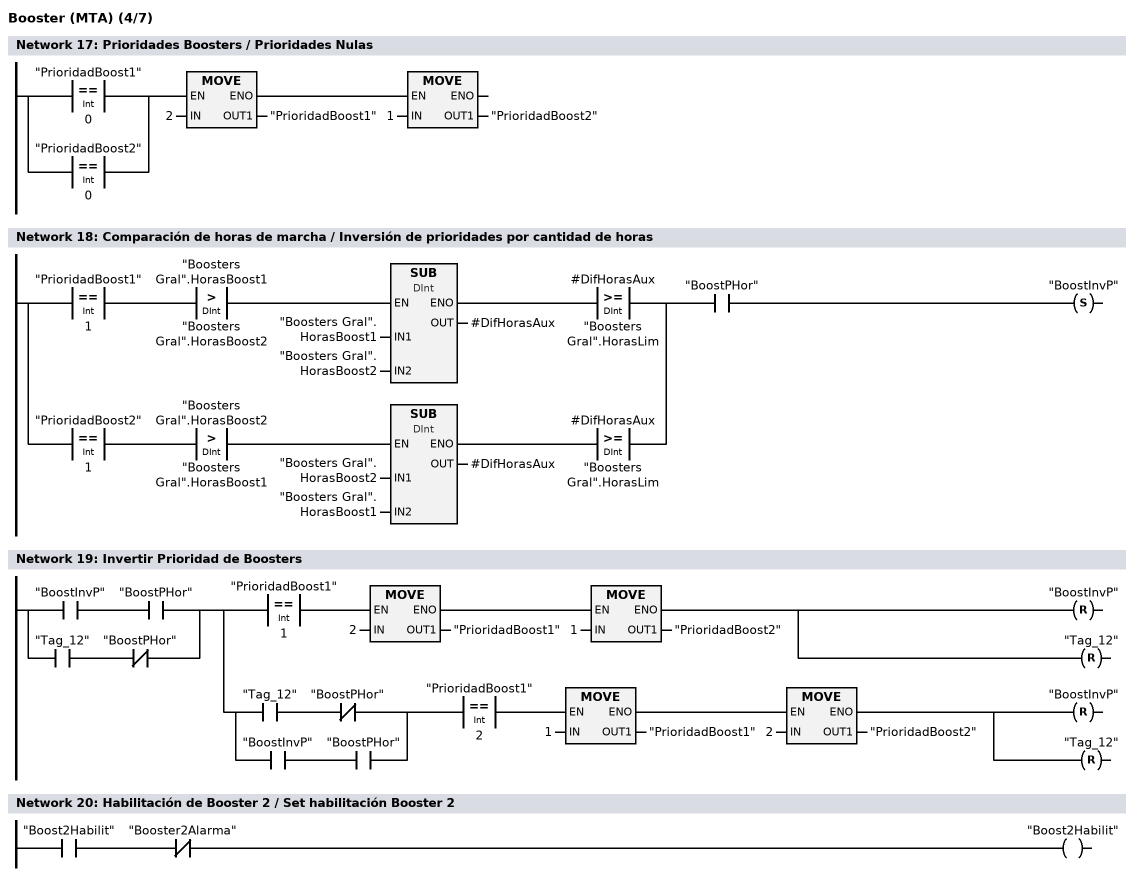
   RUNG wire#powerrail
      { S7_Templates := "SrcType := Int" } EQ_Contact(in1 := "PrioridadBoost1", in2 := 0)
      wire#w1
      { S7_GenerateENO := "TRUE" } Move(in := 2, out1 => "PrioridadBoost1")
      { S7_GenerateENO := "TRUE" } Move(in := 1, out1 => "PrioridadBoost2")
   END_RUNG
   RUNG wire#powerrail
      { S7_Templates := "SrcType := Int" } EQ_Contact(in1 := "PrioridadBoost2", in2 := 0)
   END_RUNG wire#w1
   // the same network as SCL:
   // ENO of a box is taken as its EN; it also drops when the box reports an error
   #_w1 := ("PrioridadBoost1" = 0) OR ("PrioridadBoost2" = 0);
   IF #_w1 THEN
       "PrioridadBoost1" := 2;
       "PrioridadBoost2" := 1;
   END_IF;
END_REGION

REGION Network 18: Comparación de horas de marcha / Inversión de prioridades por cantidad de horas
   RUNG wire#powerrail
      { S7_Templates := "SrcType := Int" } EQ_Contact(in1 := "PrioridadBoost1", in2 := 1)
      { S7_Templates := "SrcType := DInt" } GT_Contact(in1 := "Boosters Gral".HorasBoost1, in2 := "Boosters Gral".HorasBoost2)
      { S7_Templates := "SrcType := DInt"; S7_GenerateENO := "TRUE" } Sub(in1 := "Boosters Gral".HorasBoost1, in2 := "Boosters Gral".HorasBoost2, out => #DifHorasAux)
      { S7_Templates := "SrcType := DInt" } GE_Contact(in1 := #DifHorasAux, in2 := "Boosters Gral".HorasLim)
      wire#w1
      Contact( "BoostPHor" )
      S_Coil( "BoostInvP" )
   END_RUNG
   RUNG wire#powerrail
      { S7_Templates := "SrcType := Int" } EQ_Contact(in1 := "PrioridadBoost2", in2 := 1)
      { S7_Templates := "SrcType := DInt" } GT_Contact(in1 := "Boosters Gral".HorasBoost2, in2 := "Boosters Gral".HorasBoost1)
      { S7_Templates := "SrcType := DInt"; S7_GenerateENO := "TRUE" } Sub(in1 := "Boosters Gral".HorasBoost2, in2 := "Boosters Gral".HorasBoost1, out => #DifHorasAux)
      { S7_Templates := "SrcType := DInt" } GE_Contact(in1 := #DifHorasAux, in2 := "Boosters Gral".HorasLim)
   END_RUNG wire#w1
   // the same network as SCL:
   // ENO of a box is taken as its EN; it also drops when the box reports an error
   #_w1 := ("PrioridadBoost1" = 1) AND ("Boosters Gral".HorasBoost1 > "Boosters Gral".HorasBoost2);
   IF #_w1 THEN #DifHorasAux := "Boosters Gral".HorasBoost1 - "Boosters Gral".HorasBoost2; END_IF;
   #_w2 := ("PrioridadBoost2" = 1) AND ("Boosters Gral".HorasBoost2 > "Boosters Gral".HorasBoost1);
   #_w3 := #_w1 AND (#DifHorasAux >= "Boosters Gral".HorasLim);
   IF #_w2 THEN #DifHorasAux := "Boosters Gral".HorasBoost2 - "Boosters Gral".HorasBoost1; END_IF;
   IF (#_w3 OR (#_w2 AND (#DifHorasAux >= "Boosters Gral".HorasLim))) AND "BoostPHor" THEN
       "BoostInvP" := TRUE;
   END_IF;
END_REGION

REGION Network 19: Invertir Prioridad de Boosters
   RUNG wire#powerrail
      Contact( "BoostInvP" )
      Contact( "BoostPHor" )
      wire#w1
      { S7_Templates := "SrcType := Int" } EQ_Contact(in1 := "PrioridadBoost1", in2 := 1)
      { S7_GenerateENO := "TRUE" } Move(in := 2, out1 => "PrioridadBoost1")
      { S7_GenerateENO := "TRUE" } Move(in := 1, out1 => "PrioridadBoost2")
      wire#w2
      R_Coil( "BoostInvP" )
   END_RUNG
   RUNG wire#powerrail
      Contact( "Tag_12" )
      I_Contact( "BoostPHor" )
   END_RUNG wire#w1
   RUNG wire#w2
      R_Coil( "Tag_12" )
   END_RUNG
   RUNG wire#w1
      Contact( "Tag_12" )
      I_Contact( "BoostPHor" )
      wire#w3
      { S7_Templates := "SrcType := Int" } EQ_Contact(in1 := "PrioridadBoost1", in2 := 2)
      { S7_GenerateENO := "TRUE" } Move(in := 1, out1 => "PrioridadBoost1")
      { S7_GenerateENO := "TRUE" } Move(in := 2, out1 => "PrioridadBoost2")
      wire#w4
      R_Coil( "BoostInvP" )
   END_RUNG
   RUNG wire#w1
      Contact( "BoostInvP" )
      Contact( "BoostPHor" )
   END_RUNG wire#w3
   RUNG wire#w4
      R_Coil( "Tag_12" )
   END_RUNG
   // the same network as SCL:
   // ENO of a box is taken as its EN; it also drops when the box reports an error
   #_w1 := ("BoostInvP" AND "BoostPHor") OR ("Tag_12" AND NOT "BoostPHor");
   #_w2 := #_w1 AND ("PrioridadBoost1" = 1);
   IF #_w2 THEN
       "PrioridadBoost1" := 2;
       "PrioridadBoost2" := 1;
       "BoostInvP" := FALSE;
       "Tag_12" := FALSE;
   END_IF;
   #_w3 := #_w1 AND (("Tag_12" AND NOT "BoostPHor") OR ("BoostInvP" AND "BoostPHor")) AND ("PrioridadBoost1" = 2);
   IF #_w3 THEN
       "PrioridadBoost1" := 1;
       "PrioridadBoost2" := 2;
       "BoostInvP" := FALSE;
       "Tag_12" := FALSE;
   END_IF;
END_REGION

REGION Network 20: Habilitación de Booster 2 / Set habilitación Booster 2
   RUNG wire#powerrail
      Contact( "Boost2Habilit" )
      I_Contact( "Booster2Alarma" )
      Coil( "Boost2Habilit" )
   END_RUNG
   // the same network as SCL:
   "Boost2Habilit" := "Boost2Habilit" AND NOT "Booster2Alarma";
END_REGION

REGION Network 21: Orden de Marcha Booster
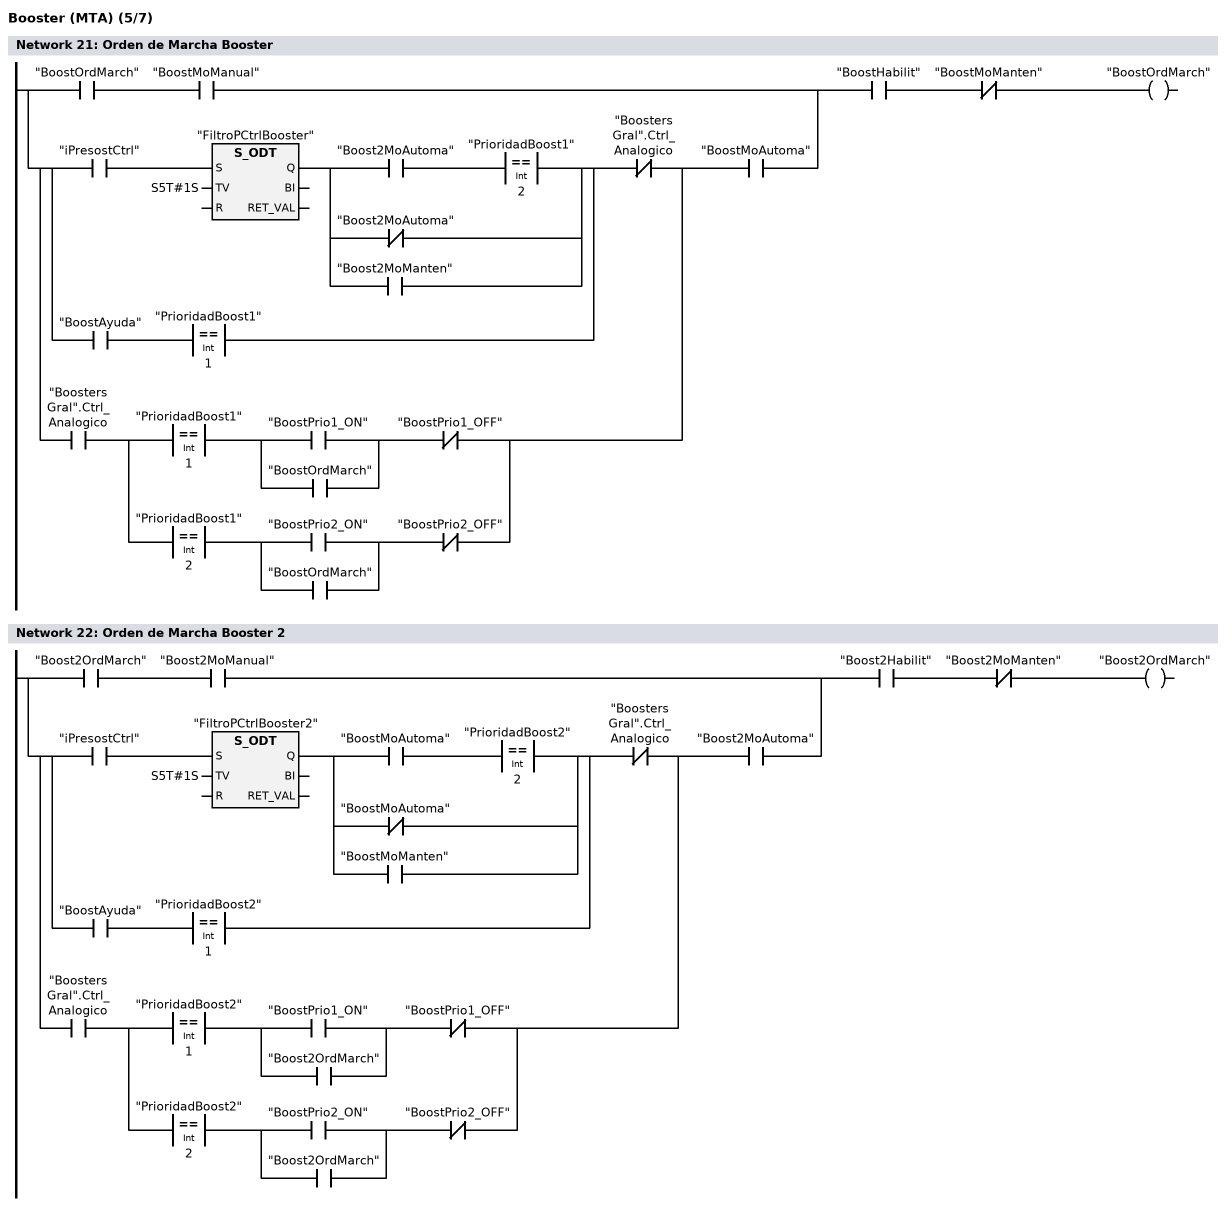
   RUNG wire#powerrail
      Contact( "BoostOrdMarch" )
      Contact( "BoostMoManual" )
      wire#w1
      Contact( "BoostHabilit" )
      I_Contact( "BoostMoManten" )
      Coil( "BoostOrdMarch" )
   END_RUNG
   RUNG wire#powerrail
      Contact( "iPresostCtrl" )
      S_ODT(T_NO := "FiltroPCtrlBooster", TV := S5T#1S, R :=, BI =>, RET_VAL =>)
      wire#w2
      Contact( "Boost2MoAutoma" )
      { S7_Templates := "SrcType := Int" } EQ_Contact(in1 := "PrioridadBoost1", in2 := 2)
      wire#w3
      I_Contact( "Boosters Gral".Ctrl_Analogico )
      wire#w4
      Contact( "BoostMoAutoma" )
   END_RUNG wire#w1
   RUNG wire#w2
      I_Contact( "Boost2MoAutoma" )
   END_RUNG wire#w3
   RUNG wire#w2
      Contact( "Boost2MoManten" )
   END_RUNG wire#w3
   RUNG wire#powerrail
      Contact( "BoostAyuda" )
      { S7_Templates := "SrcType := Int" } EQ_Contact(in1 := "PrioridadBoost1", in2 := 1)
   END_RUNG wire#w3
   RUNG wire#powerrail
      Contact( "Boosters Gral".Ctrl_Analogico )
      wire#w5
      { S7_Templates := "SrcType := Int" } EQ_Contact(in1 := "PrioridadBoost1", in2 := 1)
      wire#w6
      Contact( "BoostPrio1_ON" )
      wire#w7
      I_Contact( "BoostPrio1_OFF" )
   END_RUNG wire#w4
   RUNG wire#w6
      Contact( "BoostOrdMarch" )
   END_RUNG wire#w7
   RUNG wire#w5
      { S7_Templates := "SrcType := Int" } EQ_Contact(in1 := "PrioridadBoost1", in2 := 2)
      wire#w8
      Contact( "BoostPrio2_ON" )
      wire#w9
      I_Contact( "BoostPrio2_OFF" )
   END_RUNG wire#w4
   RUNG wire#w8
      Contact( "BoostOrdMarch" )
   END_RUNG wire#w9
   // the same network as SCL:
   #_s5time1 := S_ODT(T_NO := "FiltroPCtrlBooster", S := "iPresostCtrl", TV := S5T#1S, Q => #_w1);
   "BoostOrdMarch" := (("BoostOrdMarch" AND "BoostMoManual") OR (((((#_w1 AND (("Boost2MoAutoma" AND ("PrioridadBoost1" = 2)) OR NOT "Boost2MoAutoma" OR "Boost2MoManten")) OR ("BoostAyuda" AND ("PrioridadBoost1" = 1))) AND NOT "Boosters Gral".Ctrl_Analogico) OR ("Boosters Gral".Ctrl_Analogico AND ((("PrioridadBoost1" = 1) AND ("BoostPrio1_ON" OR "BoostOrdMarch") AND NOT "BoostPrio1_OFF") OR (("PrioridadBoost1" = 2) AND ("BoostPrio2_ON" OR "BoostOrdMarch") AND NOT "BoostPrio2_OFF")))) AND "BoostMoAutoma")) AND "BoostHabilit" AND NOT "BoostMoManten";
END_REGION

REGION Network 22: Orden de Marcha Booster 2
   RUNG wire#powerrail
      Contact( "Boost2OrdMarch" )
      Contact( "Boost2MoManual" )
      wire#w1
      Contact( "Boost2Habilit" )
      I_Contact( "Boost2MoManten" )
      Coil( "Boost2OrdMarch" )
   END_RUNG
   RUNG wire#powerrail
      Contact( "iPresostCtrl" )
      S_ODT(T_NO := "FiltroPCtrlBooster2", TV := S5T#1S, R :=, BI =>, RET_VAL =>)
      wire#w2
      Contact( "BoostMoAutoma" )
      { S7_Templates := "SrcType := Int" } EQ_Contact(in1 := "PrioridadBoost2", in2 := 2)
      wire#w3
      I_Contact( "Boosters Gral".Ctrl_Analogico )
      wire#w4
      Contact( "Boost2MoAutoma" )
   END_RUNG wire#w1
   RUNG wire#w2
      I_Contact( "BoostMoAutoma" )
   END_RUNG wire#w3
   RUNG wire#w2
      Contact( "BoostMoManten" )
   END_RUNG wire#w3
   RUNG wire#powerrail
      Contact( "BoostAyuda" )
      { S7_Templates := "SrcType := Int" } EQ_Contact(in1 := "PrioridadBoost2", in2 := 1)
   END_RUNG wire#w3
   RUNG wire#powerrail
      Contact( "Boosters Gral".Ctrl_Analogico )
      wire#w5
      { S7_Templates := "SrcType := Int" } EQ_Contact(in1 := "PrioridadBoost2", in2 := 1)
      wire#w6
      Contact( "BoostPrio1_ON" )
      wire#w7
      I_Contact( "BoostPrio1_OFF" )
   END_RUNG wire#w4
   RUNG wire#w6
      Contact( "Boost2OrdMarch" )
   END_RUNG wire#w7
   RUNG wire#w5
      { S7_Templates := "SrcType := Int" } EQ_Contact(in1 := "PrioridadBoost2", in2 := 2)
      wire#w8
      Contact( "BoostPrio2_ON" )
      wire#w9
      I_Contact( "BoostPrio2_OFF" )
   END_RUNG wire#w4
   RUNG wire#w8
      Contact( "Boost2OrdMarch" )
   END_RUNG wire#w9
   // the same network as SCL:
   #_s5time1 := S_ODT(T_NO := "FiltroPCtrlBooster2", S := "iPresostCtrl", TV := S5T#1S, Q => #_w1);
   "Boost2OrdMarch" := (("Boost2OrdMarch" AND "Boost2MoManual") OR (((((#_w1 AND (("BoostMoAutoma" AND ("PrioridadBoost2" = 2)) OR NOT "BoostMoAutoma" OR "BoostMoManten")) OR ("BoostAyuda" AND ("PrioridadBoost2" = 1))) AND NOT "Boosters Gral".Ctrl_Analogico) OR ("Boosters Gral".Ctrl_Analogico AND ((("PrioridadBoost2" = 1) AND ("BoostPrio1_ON" OR "Boost2OrdMarch") AND NOT "BoostPrio1_OFF") OR (("PrioridadBoost2" = 2) AND ("BoostPrio2_ON" OR "Boost2OrdMarch") AND NOT "BoostPrio2_OFF")))) AND "Boost2MoAutoma")) AND "Boost2Habilit" AND NOT "Boost2MoManten";
END_REGION

REGION Network 23: Motor Booster 1 / Bloque de Motor Booster
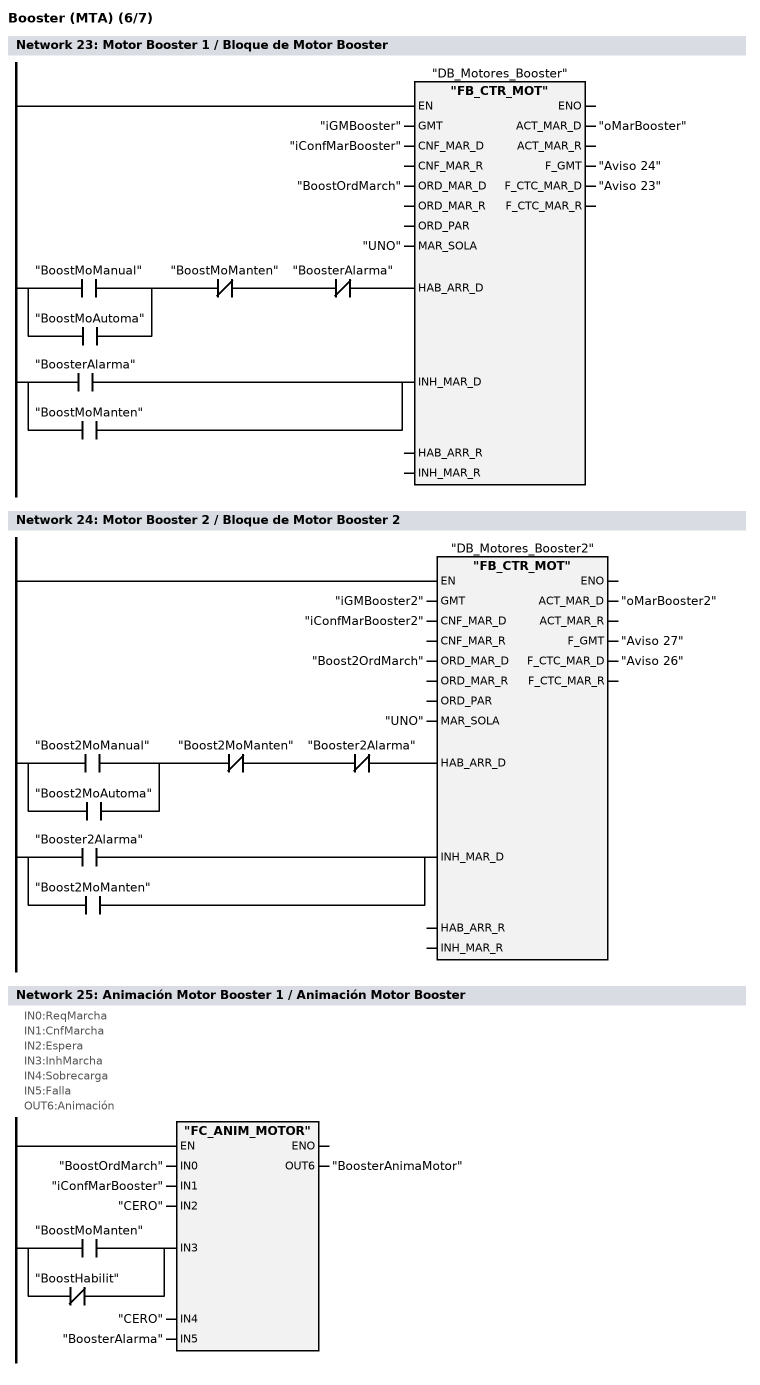
   RUNG wire#powerrail
      "DB_Motores_Booster"(HAB_ARR_D := wire#w2, INH_MAR_D := wire#w3, GMT := "iGMBooster", CNF_MAR_D := "iConfMarBooster", CNF_MAR_R :=, ORD_MAR_D := "BoostOrdMarch", ORD_MAR_R :=, ORD_PAR :=, MAR_SOLA := "UNO", HAB_ARR_R :=, INH_MAR_R :=, ACT_MAR_D => "oMarBooster", ACT_MAR_R =>, F_GMT => "Aviso 24", F_CTC_MAR_D => "Aviso 23", F_CTC_MAR_R =>)
   END_RUNG
   RUNG wire#powerrail
      Contact( "BoostMoManual" )
      wire#w1
      I_Contact( "BoostMoManten" )
      I_Contact( "BoosterAlarma" )
   END_RUNG wire#w2
   RUNG wire#powerrail
      Contact( "BoostMoAutoma" )
   END_RUNG wire#w1
   RUNG wire#powerrail
      Contact( "BoosterAlarma" )
   END_RUNG wire#w3
   RUNG wire#powerrail
      Contact( "BoostMoManten" )
   END_RUNG wire#w3
   // the same network as SCL:
   "DB_Motores_Booster"(GMT := "iGMBooster",   // "FB_CTR_MOT"
                        CNF_MAR_D := "iConfMarBooster",
                        ORD_MAR_D := "BoostOrdMarch",
                        MAR_SOLA := "UNO",
                        HAB_ARR_D := ("BoostMoManual" OR "BoostMoAutoma") AND NOT "BoostMoManten" AND NOT "BoosterAlarma",
                        INH_MAR_D := "BoosterAlarma" OR "BoostMoManten",
                        ACT_MAR_D => "oMarBooster",
                        F_GMT => "Aviso 24",
                        F_CTC_MAR_D => "Aviso 23");
END_REGION

REGION Network 24: Motor Booster 2 / Bloque de Motor Booster 2
   RUNG wire#powerrail
      "DB_Motores_Booster2"(HAB_ARR_D := wire#w2, INH_MAR_D := wire#w3, GMT := "iGMBooster2", CNF_MAR_D := "iConfMarBooster2", CNF_MAR_R :=, ORD_MAR_D := "Boost2OrdMarch", ORD_MAR_R :=, ORD_PAR :=, MAR_SOLA := "UNO", HAB_ARR_R :=, INH_MAR_R :=, ACT_MAR_D => "oMarBooster2", ACT_MAR_R =>, F_GMT => "Aviso 27", F_CTC_MAR_D => "Aviso 26", F_CTC_MAR_R =>)
   END_RUNG
   RUNG wire#powerrail
      Contact( "Boost2MoManual" )
      wire#w1
      I_Contact( "Boost2MoManten" )
      I_Contact( "Booster2Alarma" )
   END_RUNG wire#w2
   RUNG wire#powerrail
      Contact( "Boost2MoAutoma" )
   END_RUNG wire#w1
   RUNG wire#powerrail
      Contact( "Booster2Alarma" )
   END_RUNG wire#w3
   RUNG wire#powerrail
      Contact( "Boost2MoManten" )
   END_RUNG wire#w3
   // the same network as SCL:
   "DB_Motores_Booster2"(GMT := "iGMBooster2",   // "FB_CTR_MOT"
                         CNF_MAR_D := "iConfMarBooster2",
                         ORD_MAR_D := "Boost2OrdMarch",
                         MAR_SOLA := "UNO",
                         HAB_ARR_D := ("Boost2MoManual" OR "Boost2MoAutoma") AND NOT "Boost2MoManten" AND NOT "Booster2Alarma",
                         INH_MAR_D := "Booster2Alarma" OR "Boost2MoManten",
                         ACT_MAR_D => "oMarBooster2",
                         F_GMT => "Aviso 27",
                         F_CTC_MAR_D => "Aviso 26");
END_REGION

REGION Network 25: Animación Motor Booster 1 / Animación Motor Booster
   // IN0:ReqMarcha
   // IN1:CnfMarcha
   // IN2:Espera
   // IN3:InhMarcha
   // IN4:Sobrecarga
   // IN5:Falla
   // OUT6:Animación
   RUNG wire#powerrail
      "FC_ANIM_MOTOR"(IN0 := "BoostOrdMarch", IN1 := "iConfMarBooster", IN2 := "CERO", IN3 := wire#w1, IN4 := "CERO", IN5 := "BoosterAlarma", OUT6 => "BoosterAnimaMotor")
   END_RUNG
   RUNG wire#powerrail
      Contact( "BoostMoManten" )
   END_RUNG wire#w1
   RUNG wire#powerrail
      I_Contact( "BoostHabilit" )
   END_RUNG wire#w1
   // the same network as SCL:
   "FC_ANIM_MOTOR"(IN0 := "BoostOrdMarch",
                   IN1 := "iConfMarBooster",
                   IN2 := "CERO",
                   IN3 := "BoostMoManten" OR NOT "BoostHabilit",
                   IN4 := "CERO",
                   IN5 := "BoosterAlarma",
                   OUT6 => "BoosterAnimaMotor");
END_REGION

REGION Network 26: Animación Motor Booster 2
   // IN0:ReqMarcha
   // IN1:CnfMarcha
   // IN2:Espera
   // IN3:InhMarcha
   // IN4:Sobrecarga
   // IN5:Falla
   // OUT6:Animación
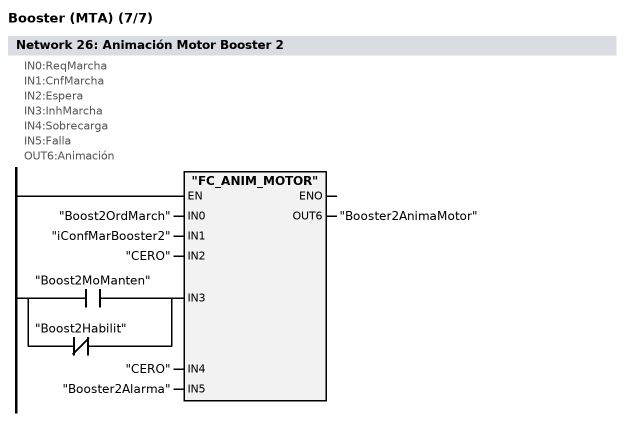
   RUNG wire#powerrail
      "FC_ANIM_MOTOR"(IN0 := "Boost2OrdMarch", IN1 := "iConfMarBooster2", IN2 := "CERO", IN3 := wire#w1, IN4 := "CERO", IN5 := "Booster2Alarma", OUT6 => "Booster2AnimaMotor")
   END_RUNG
   RUNG wire#powerrail
      Contact( "Boost2MoManten" )
   END_RUNG wire#w1
   RUNG wire#powerrail
      I_Contact( "Boost2Habilit" )
   END_RUNG wire#w1
   // the same network as SCL:
   "FC_ANIM_MOTOR"(IN0 := "Boost2OrdMarch",
                   IN1 := "iConfMarBooster2",
                   IN2 := "CERO",
                   IN3 := "Boost2MoManten" OR NOT "Boost2Habilit",
                   IN4 := "CERO",
                   IN5 := "Booster2Alarma",
                   OUT6 => "Booster2AnimaMotor");
END_REGION
END_FUNCTION

// folder: Compresores/Alta

FUNCTION "CompresoresAltaMTA" : Void   // FC13, LAD
{ S7_Optimized_Access := 'FALSE' }
VERSION : 0.1
BEGIN

REGION Network 1
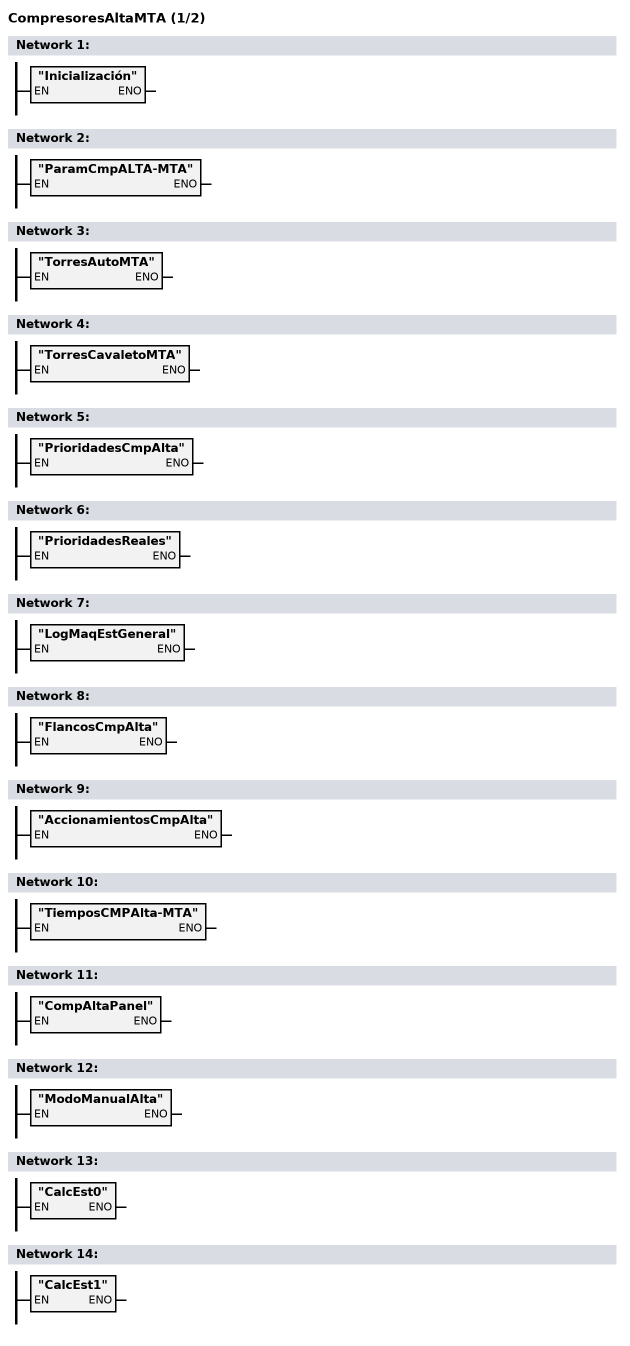
   RUNG wire#powerrail
      "Inicialización"()
   END_RUNG
   // the same network as SCL:
   "Inicialización"();
END_REGION

REGION Network 2
   RUNG wire#powerrail
      "ParamCmpALTA-MTA"()
   END_RUNG
   // the same network as SCL:
   "ParamCmpALTA-MTA"();
END_REGION

REGION Network 3
   RUNG wire#powerrail
      "TorresAutoMTA"()
   END_RUNG
   // the same network as SCL:
   "TorresAutoMTA"();
END_REGION

REGION Network 4
   RUNG wire#powerrail
      "TorresCavaletoMTA"()
   END_RUNG
   // the same network as SCL:
   "TorresCavaletoMTA"();
END_REGION

REGION Network 5
   RUNG wire#powerrail
      "PrioridadesCmpAlta"()
   END_RUNG
   // the same network as SCL:
   "PrioridadesCmpAlta"();
END_REGION

REGION Network 6
   RUNG wire#powerrail
      "PrioridadesReales"()
   END_RUNG
   // the same network as SCL:
   "PrioridadesReales"();
END_REGION

REGION Network 7
   RUNG wire#powerrail
      "LogMaqEstGeneral"()
   END_RUNG
   // the same network as SCL:
   "LogMaqEstGeneral"();
END_REGION

REGION Network 8
   RUNG wire#powerrail
      "FlancosCmpAlta"()
   END_RUNG
   // the same network as SCL:
   "FlancosCmpAlta"();
END_REGION

REGION Network 9
   RUNG wire#powerrail
      "AccionamientosCmpAlta"()
   END_RUNG
   // the same network as SCL:
   "AccionamientosCmpAlta"();
END_REGION

REGION Network 10
   RUNG wire#powerrail
      "TiemposCMPAlta-MTA"()
   END_RUNG
   // the same network as SCL:
   "TiemposCMPAlta-MTA"();
END_REGION

REGION Network 11
   RUNG wire#powerrail
      "CompAltaPanel"()
   END_RUNG
   // the same network as SCL:
   "CompAltaPanel"();
END_REGION

REGION Network 12
   RUNG wire#powerrail
      "ModoManualAlta"()
   END_RUNG
   // the same network as SCL:
   "ModoManualAlta"();
END_REGION

REGION Network 13
   RUNG wire#powerrail
      "CalcEst0"()
   END_RUNG
   // the same network as SCL:
   "CalcEst0"();
END_REGION

REGION Network 14
   RUNG wire#powerrail
      "CalcEst1"()
   END_RUNG
   // the same network as SCL:
   "CalcEst1"();
END_REGION

REGION Network 15
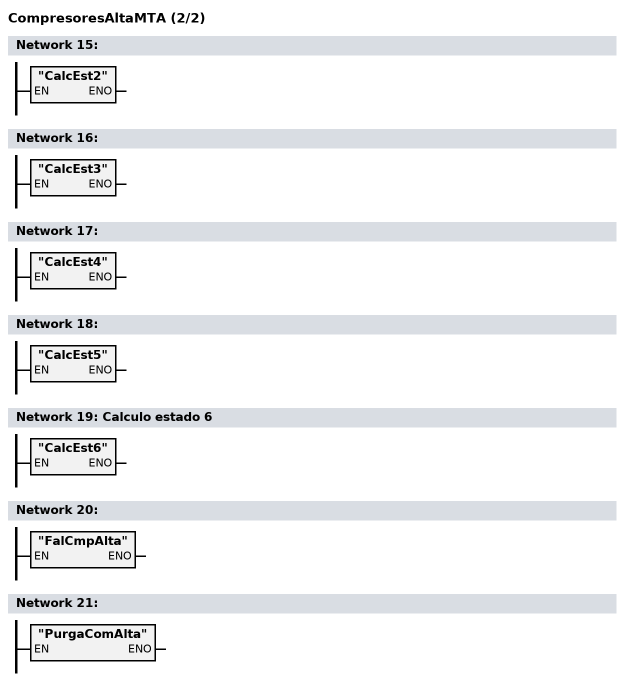
   RUNG wire#powerrail
      "CalcEst2"()
   END_RUNG
   // the same network as SCL:
   "CalcEst2"();
END_REGION

REGION Network 16
   RUNG wire#powerrail
      "CalcEst3"()
   END_RUNG
   // the same network as SCL:
   "CalcEst3"();
END_REGION

REGION Network 17
   RUNG wire#powerrail
      "CalcEst4"()
   END_RUNG
   // the same network as SCL:
   "CalcEst4"();
END_REGION

REGION Network 18
   RUNG wire#powerrail
      "CalcEst5"()
   END_RUNG
   // the same network as SCL:
   "CalcEst5"();
END_REGION

REGION Network 19: Calculo estado 6
   RUNG wire#powerrail
      "CalcEst6"()
   END_RUNG
   // the same network as SCL:
   "CalcEst6"();
END_REGION

REGION Network 20
   RUNG wire#powerrail
      "FalCmpAlta"()
   END_RUNG
   // the same network as SCL:
   "FalCmpAlta"();
END_REGION

REGION Network 21
   RUNG wire#powerrail
      "PurgaComAlta"()
   END_RUNG
   // the same network as SCL:
   "PurgaComAlta"();
END_REGION
END_FUNCTION

FUNCTION "ParamCmpALTA-MTA" : Void   // FC30, LAD
{ S7_Optimized_Access := 'FALSE' }
VERSION : 0.1
BEGIN

REGION Network 1
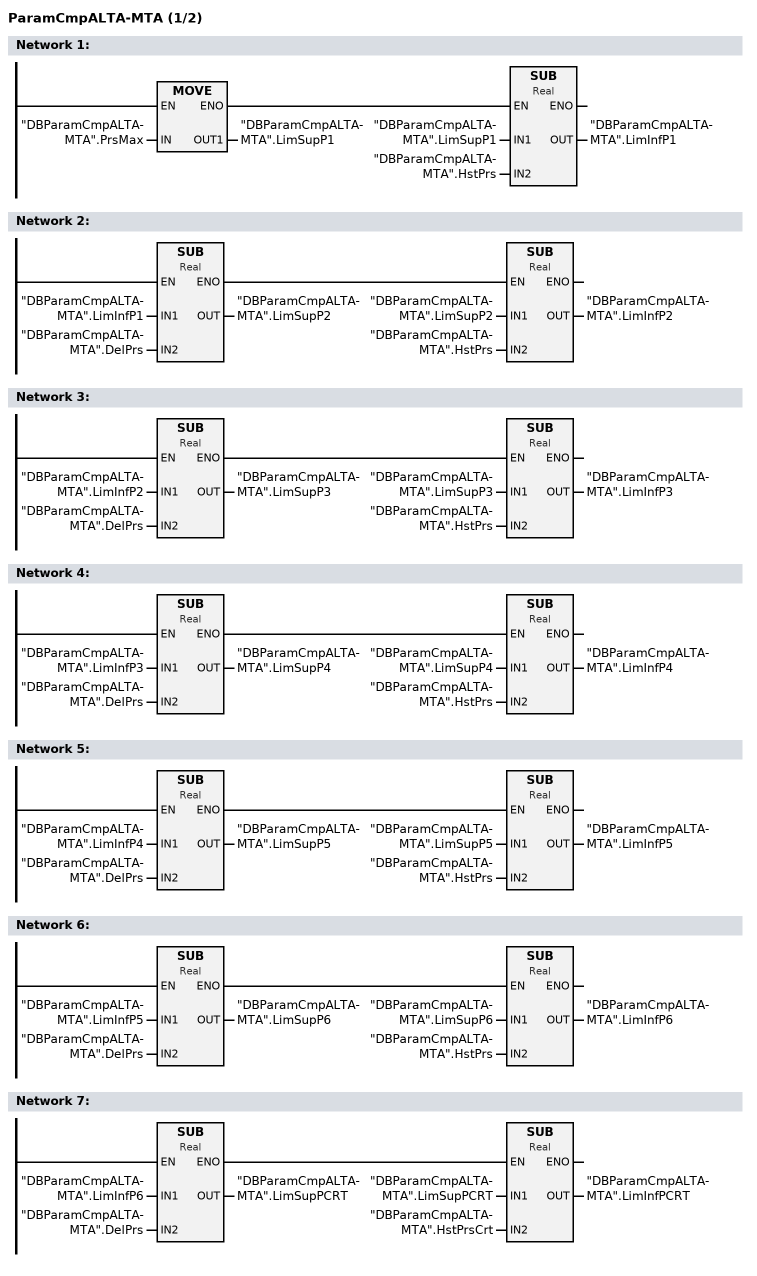
   RUNG wire#powerrail
      { S7_GenerateENO := "TRUE" } Move(in := "DBParamCmpALTA-MTA".PrsMax, out1 => "DBParamCmpALTA-MTA".LimSupP1)
      { S7_Templates := "SrcType := Real"; S7_GenerateENO := "TRUE" } Sub(in1 := "DBParamCmpALTA-MTA".LimSupP1, in2 := "DBParamCmpALTA-MTA".HstPrs, out => "DBParamCmpALTA-MTA".LimInfP1)
   END_RUNG
   // the same network as SCL:
   // ENO of a box is taken as its EN; it also drops when the box reports an error
   "DBParamCmpALTA-MTA".LimSupP1 := "DBParamCmpALTA-MTA".PrsMax;
   "DBParamCmpALTA-MTA".LimInfP1 := "DBParamCmpALTA-MTA".LimSupP1 - "DBParamCmpALTA-MTA".HstPrs;
END_REGION

REGION Network 2
   RUNG wire#powerrail
      { S7_Templates := "SrcType := Real"; S7_GenerateENO := "TRUE" } Sub(in1 := "DBParamCmpALTA-MTA".LimInfP1, in2 := "DBParamCmpALTA-MTA".DelPrs, out => "DBParamCmpALTA-MTA".LimSupP2)
      { S7_Templates := "SrcType := Real"; S7_GenerateENO := "TRUE" } Sub(in1 := "DBParamCmpALTA-MTA".LimSupP2, in2 := "DBParamCmpALTA-MTA".HstPrs, out => "DBParamCmpALTA-MTA".LimInfP2)
   END_RUNG
   // the same network as SCL:
   // ENO of a box is taken as its EN; it also drops when the box reports an error
   "DBParamCmpALTA-MTA".LimSupP2 := "DBParamCmpALTA-MTA".LimInfP1 - "DBParamCmpALTA-MTA".DelPrs;
   "DBParamCmpALTA-MTA".LimInfP2 := "DBParamCmpALTA-MTA".LimSupP2 - "DBParamCmpALTA-MTA".HstPrs;
END_REGION

REGION Network 3
   RUNG wire#powerrail
      { S7_Templates := "SrcType := Real"; S7_GenerateENO := "TRUE" } Sub(in1 := "DBParamCmpALTA-MTA".LimInfP2, in2 := "DBParamCmpALTA-MTA".DelPrs, out => "DBParamCmpALTA-MTA".LimSupP3)
      { S7_Templates := "SrcType := Real"; S7_GenerateENO := "TRUE" } Sub(in1 := "DBParamCmpALTA-MTA".LimSupP3, in2 := "DBParamCmpALTA-MTA".HstPrs, out => "DBParamCmpALTA-MTA".LimInfP3)
   END_RUNG
   // the same network as SCL:
   // ENO of a box is taken as its EN; it also drops when the box reports an error
   "DBParamCmpALTA-MTA".LimSupP3 := "DBParamCmpALTA-MTA".LimInfP2 - "DBParamCmpALTA-MTA".DelPrs;
   "DBParamCmpALTA-MTA".LimInfP3 := "DBParamCmpALTA-MTA".LimSupP3 - "DBParamCmpALTA-MTA".HstPrs;
END_REGION

REGION Network 4
   RUNG wire#powerrail
      { S7_Templates := "SrcType := Real"; S7_GenerateENO := "TRUE" } Sub(in1 := "DBParamCmpALTA-MTA".LimInfP3, in2 := "DBParamCmpALTA-MTA".DelPrs, out => "DBParamCmpALTA-MTA".LimSupP4)
      { S7_Templates := "SrcType := Real"; S7_GenerateENO := "TRUE" } Sub(in1 := "DBParamCmpALTA-MTA".LimSupP4, in2 := "DBParamCmpALTA-MTA".HstPrs, out => "DBParamCmpALTA-MTA".LimInfP4)
   END_RUNG
   // the same network as SCL:
   // ENO of a box is taken as its EN; it also drops when the box reports an error
   "DBParamCmpALTA-MTA".LimSupP4 := "DBParamCmpALTA-MTA".LimInfP3 - "DBParamCmpALTA-MTA".DelPrs;
   "DBParamCmpALTA-MTA".LimInfP4 := "DBParamCmpALTA-MTA".LimSupP4 - "DBParamCmpALTA-MTA".HstPrs;
END_REGION

REGION Network 5
   RUNG wire#powerrail
      { S7_Templates := "SrcType := Real"; S7_GenerateENO := "TRUE" } Sub(in1 := "DBParamCmpALTA-MTA".LimInfP4, in2 := "DBParamCmpALTA-MTA".DelPrs, out => "DBParamCmpALTA-MTA".LimSupP5)
      { S7_Templates := "SrcType := Real"; S7_GenerateENO := "TRUE" } Sub(in1 := "DBParamCmpALTA-MTA".LimSupP5, in2 := "DBParamCmpALTA-MTA".HstPrs, out => "DBParamCmpALTA-MTA".LimInfP5)
   END_RUNG
   // the same network as SCL:
   // ENO of a box is taken as its EN; it also drops when the box reports an error
   "DBParamCmpALTA-MTA".LimSupP5 := "DBParamCmpALTA-MTA".LimInfP4 - "DBParamCmpALTA-MTA".DelPrs;
   "DBParamCmpALTA-MTA".LimInfP5 := "DBParamCmpALTA-MTA".LimSupP5 - "DBParamCmpALTA-MTA".HstPrs;
END_REGION

REGION Network 6
   RUNG wire#powerrail
      { S7_Templates := "SrcType := Real"; S7_GenerateENO := "TRUE" } Sub(in1 := "DBParamCmpALTA-MTA".LimInfP5, in2 := "DBParamCmpALTA-MTA".DelPrs, out => "DBParamCmpALTA-MTA".LimSupP6)
      { S7_Templates := "SrcType := Real"; S7_GenerateENO := "TRUE" } Sub(in1 := "DBParamCmpALTA-MTA".LimSupP6, in2 := "DBParamCmpALTA-MTA".HstPrs, out => "DBParamCmpALTA-MTA".LimInfP6)
   END_RUNG
   // the same network as SCL:
   // ENO of a box is taken as its EN; it also drops when the box reports an error
   "DBParamCmpALTA-MTA".LimSupP6 := "DBParamCmpALTA-MTA".LimInfP5 - "DBParamCmpALTA-MTA".DelPrs;
   "DBParamCmpALTA-MTA".LimInfP6 := "DBParamCmpALTA-MTA".LimSupP6 - "DBParamCmpALTA-MTA".HstPrs;
END_REGION

REGION Network 7
   RUNG wire#powerrail
      { S7_Templates := "SrcType := Real"; S7_GenerateENO := "TRUE" } Sub(in1 := "DBParamCmpALTA-MTA".LimInfP6, in2 := "DBParamCmpALTA-MTA".DelPrs, out => "DBParamCmpALTA-MTA".LimSupPCRT)
      { S7_Templates := "SrcType := Real"; S7_GenerateENO := "TRUE" } Sub(in1 := "DBParamCmpALTA-MTA".LimSupPCRT, in2 := "DBParamCmpALTA-MTA".HstPrsCrt, out => "DBParamCmpALTA-MTA".LimInfPCRT)
   END_RUNG
   // the same network as SCL:
   // ENO of a box is taken as its EN; it also drops when the box reports an error
   "DBParamCmpALTA-MTA".LimSupPCRT := "DBParamCmpALTA-MTA".LimInfP6 - "DBParamCmpALTA-MTA".DelPrs;
   "DBParamCmpALTA-MTA".LimInfPCRT := "DBParamCmpALTA-MTA".LimSupPCRT - "DBParamCmpALTA-MTA".HstPrsCrt;
END_REGION

REGION Network 8: Falla General Flujostato Cavaleto
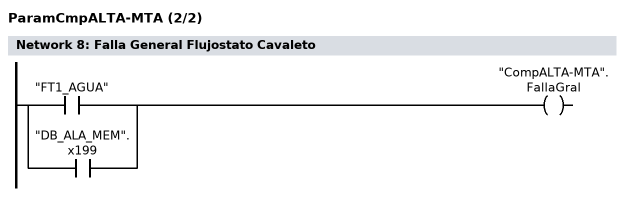
   RUNG wire#powerrail
      Contact( "FT1_AGUA" )
      wire#w1
      Coil( "CompALTA-MTA".FallaGral )
   END_RUNG
   RUNG wire#powerrail
      Contact( "DB_ALA_MEM".x199 )
   END_RUNG wire#w1
   // the same network as SCL:
   "CompALTA-MTA".FallaGral := "FT1_AGUA" OR "DB_ALA_MEM".x199;
END_REGION
END_FUNCTION

FUNCTION "TiemposCMPAlta-MTA" : Void   // FC31, LAD
{ S7_Optimized_Access := 'FALSE' }
VERSION : 0.1
   VAR_TEMP   // added for the SCL form of the ladder/FBD networks
      _s5time1 : S5Time;
   END_VAR
BEGIN

REGION Network 1